HMI tags "AO"
   "DB332_AO_AO{1}_bRoZB1" : Byte = PLC DB332_AO.AO[1].bRoZB1, 1 s
   "DB332_AO_AO{1}_bSym" : Word = PLC DB332_AO.AO[1].bSym AT %DB1.DBB0, 1 s
   "DB332_AO_AO{1}_bSt_Tryb" : Word = PLC DB332_AO.AO[1].bSt_Tryb AT %DB1.DBW0, 1 s
   "DB332_AO_AO{1}_bSt_Urz" : Int = PLC DB332_AO.AO[1].bSt_Urz, 1 s
   "DB332_AO_AO{1}_bTrP" : Int = PLC DB332_AO.AO[1].bTrP AT %DB1.DBW0, 1 s
   "DB332_AO_AO{1}_yCzZadFiltru" : Byte = PLC DB332_AO.AO[1].yCzZadFiltru AT %DB1.DBW0, 1 s
   "DB332_AO_AO{1}_bB" : Byte = PLC DB332_AO.AO[1].bB AT %DB1.DBW0, 1 s
   "DB332_AO_AO{1}_rZH" : Real = PLC DB332_AO.AO[1].rZH AT %DB1.DBB0, 1 s
   "DB332_AO_AO{Nr}_rZL" : Real = PLC DB332_AO.AO[1].rZL AT %DB1.DBD0, 1 s
   "DB332_AO_AO{Nr}_rGHH" : Real = PLC DB332_AO.AO[1].rGHH AT %DB1.DBD0, 1 s
   "DB332_AO_AO{Nr}_rGH" : Real = PLC DB332_AO.AO[1].rGH AT %DB1.DBD0, 1 s
   "DB332_AO_AO{Nr}_rGL" : Real = PLC DB332_AO.AO[1].rGL AT %DB1.DBD0, 1 s
   "DB332_AO_AO{Nr}_rGLL" : Real = PLC DB332_AO.AO[1].rGLL AT %DB1.DBD0, 1 s
   "DB332_AO_AO{Nr}_rHI_LIM" : Real = PLC DB332_AO.AO[1].rHI_LIM, 1 s
   "DB332_AO_AO{Nr}_rRoManSter" : Real = PLC DB332_AO.AO[1].rRoManSter, 1 s
   "DB332_AO_AO{Nr}_rWy" : Real = PLC DB332_AO.AO[1].rWy, 1 s

HMI tags "DIO"
   "DB321_DIO_DIO{Nr}_bRoZB1" : Byte = PLC DB321_DIO.DIO[1].bRoZB1, 1 s
   "DB321_DIO_DIO{Nr}_bSt_Tryb" : Word = PLC DB321_DIO.DIO[1].bSt_Tryb AT %DB1.DBB0, 1 s
   "DB321_DIO_DIO{Nr}_bWySter" : Bool = PLC DB321_DIO.DIO[1].bWySter AT %DB1.DBW0, 1 s
   "DB321_DIO_DIO{Nr}_yCzZadOpzZal" : DWord = PLC DB321_DIO.DIO[1].yCzZadOpzZal AT %DB1.DBX0.0, 1 s
   "DB321_DIO_DIO{Nr}_yCzZadOpzWyl" : DWord = PLC DB321_DIO.DIO[1].yCzZadOpzWyl AT %DB1.DBD0, 1 s

HMI tags "DM"
   "DB323_DM1_DM1{Nr}_bRoZB1" : Byte = PLC DB323_DM1.DM1[1].bRoZB1, 1 s
   "DB323_DM1_DM1{Nr}_bRoZB2" : Byte = PLC DB323_DM1.DM1[1].bRoZB2 AT %DB1.DBB0, 1 s
   "DB323_DM1_DM1{Nr}_bSym" : Word = PLC DB323_DM1.DM1[1].bSym AT %DB1.DBB0, 1 s
   "DB323_DM1_DM1{Nr}_bSt_Tryb" : Word = PLC DB323_DM1.DM1[1].bSt_Tryb AT %DB1.DBW0, 1 s
   "DB323_DM1_DM1{Nr}_bSt_Urz" : Int = PLC DB323_DM1.DM1[1].bSt_Urz AT %DB1.DBW0, 1 s
   "DB323_DM1_DM1{Nr}_bTrP" : Int = PLC DB323_DM1.DM1[1].bTrP AT %DB1.DBW0, 1 s
   "DB323_DM1_DM1{Nr}_yCzZadOpzZal" : DWord = PLC DB323_DM1.DM1[1].yCzZadOpzZal AT %DB1.DBW0, 1 s
   "DB323_DM1_DM1{Nr}_yCzZadOpzWyl" : DWord = PLC DB323_DM1.DM1[1].yCzZadOpzWyl AT %DB1.DBD0, 1 s
   "DB323_DM1_DM1{1}" : UDT323_DM1 = PLC DB323_DM1.DM1[1] AT %DB1.DBB0, 1 s
   "DB323_DM1_DM1{2}" : UDT323_DM1 = PLC DB323_DM1.DM1[2] AT %DB1.DBW0, 1 s
   "DB323_DM1_DM1{3}" : UDT323_DM1 = PLC DB323_DM1.DM1[3] AT %DB1.DBW0, 1 s
   "DB323_DM1_DM1{4}" : UDT323_DM1 = PLC DB323_DM1.DM1[4] AT %DB1.DBW0, 1 s
   "DB323_DM1_DM1{5}" : UDT323_DM1 = PLC DB323_DM1.DM1[5] AT %DB1.DBW0, 1 s
   "DB323_DM1_DM1{Nr}_yCzZadOpzAlm" : Byte = PLC DB323_DM1.DM1[1].yCzZadOpzAlm AT %DB1.DBD0, 1 s
   "DB323_DM1_DM1{Nr}_bWySter" : Bool = PLC DB323_DM1.DM1[1].bWySter AT %DB1.DBD0, 1 s

HMI tags "DV"
   "DB322_DV1_DV1{Nr}_bRoZB1" : Byte = PLC DB322_DV1.DV1[1].bRoZB1, 1 s
   "DB322_DV1_DV1{Nr}_bRoZB2" : Byte = PLC DB322_DV1.DV1[1].bRoZB2 AT %DB1.DBB0, 1 s
   "DB322_DV1_DV1{Nr}_bSym" : Word = PLC DB322_DV1.DV1[1].bSym AT %DB1.DBB0, 1 s
   "DB322_DV1_DV1{Nr}_bSt_Tryb" : Word = PLC DB322_DV1.DV1[1].bSt_Tryb AT %DB1.DBW0, 1 s
   "DB322_DV1_DV1{Nr}_bSt_Urz" : Int = PLC DB322_DV1.DV1[1].bSt_Urz AT %DB1.DBW0, 1 s
   "DB322_DV1_DV1{Nr}_bTrP" : Int = PLC DB322_DV1.DV1[1].bTrP AT %DB1.DBW0, 1 s
   "DB322_DV1_DV1{Nr}_yCzZadOpzZal" : DWord = PLC DB322_DV1.DV1[1].yCzZadOpzZal AT %DB1.DBW0, 1 s
   "DB322_DV1_DV1{Nr}_yCzZadOpzWyl" : DWord = PLC DB322_DV1.DV1[1].yCzZadOpzWyl, 1 s
   "DB322_DV1_DV1{Nr}_yCzZadOpzAlm" : Byte = PLC DB322_DV1.DV1[1].yCzZadOpzAlm AT %DB1.DBD0, 1 s
   "DB322_DV1_DV1{1}" : UDT322_DVI = PLC DB322_DV1.DV1[1] AT %DB1.DBD0, 1 s
   "DB322_DV1_DV1{2}" : UDT322_DVI = PLC DB322_DV1.DV1[2] AT %DB1.DBW0, 1 s
   "DB322_DV1_DV1{Nr}_bWySter" : Bool = PLC DB322_DV1.DV1[1].bWySter AT %DB1.DBD0, 1 s

HMI tags "Tag table_1"
   "DB_DM_pump1Tank1out_inTurnOnDelay" : DInt = PLC DB_DM.pump1Tank1out.inTurnOnDelay, 1 s
   "DB_DM_pump1Tank1out_inTurnOffDelay" : DInt = PLC DB_DM.pump1Tank1out.inTurnOffDelay, 1 s
   "DB_DM_pump1Tank1out_inAlarmDelay" : DInt = PLC DB_DM.pump1Tank1out.inAlarmDelay, 1 s
   "DB_DM_pump1Tank1out_oFaultCode" : Byte = PLC DB_DM.pump1Tank1out.oFaultCode, 1 s
   "DB_DM_pump1Tank1out_oStatusCode" : Word = PLC DB_DM.pump1Tank1out.oStatusCode, 1 s
   "DB_DM_pump1Tank1out_oStatus" : Int = PLC DB_DM.pump1Tank1out.oStatus, 1 s
   "DB_DM_pump1Tank1out_oControlMode" : Int = PLC DB_DM.pump1Tank1out.oControlMode, 1 s
   "DB_DM_pump1Tank1out_inCmdOper" : Word = PLC DB_DM.pump1Tank1out.inCmdOper, 1 s
   "DB_DM_pump1Tank1out_inSimOper" : Word = PLC DB_DM.pump1Tank1out.inSimOper, 1 s
   "DB_DM_pump1Tank1out_inCmdOperImp" : Word = PLC DB_DM.pump1Tank1out.inCmdOperImp, 1 s
   "DB_DM_pump2Tank1in_inTurnOnDelay" : DInt = PLC DB_DM.pump2Tank1in.inTurnOnDelay, 1 s
   "DB_DM_pump2Tank1in_inTurnOffDelay" : DInt = PLC DB_DM.pump2Tank1in.inTurnOffDelay, 1 s
   "DB_DM_pump2Tank1in_inAlarmDelay" : DInt = PLC DB_DM.pump2Tank1in.inAlarmDelay, 1 s
   "DB_DM_pump2Tank1in_oFaultCode" : Byte = PLC DB_DM.pump2Tank1in.oFaultCode, 1 s
   "DB_DM_pump2Tank1in_oStatusCode" : Word = PLC DB_DM.pump2Tank1in.oStatusCode, 1 s
   "DB_DM_pump2Tank1in_oStatus" : Int = PLC DB_DM.pump2Tank1in.oStatus, 1 s
   "DB_DM_pump2Tank1in_oControlMode" : Int = PLC DB_DM.pump2Tank1in.oControlMode, 1 s
   "DB_DM_pump2Tank1in_inCmdOper" : Word = PLC DB_DM.pump2Tank1in.inCmdOper, 1 s
   "DB_DM_pump2Tank1in_inSimOper" : Word = PLC DB_DM.pump2Tank1in.inSimOper, 1 s
   "DB_DM_pump2Tank1in_inCmdOperImp" : Word = PLC DB_DM.pump2Tank1in.inCmdOperImp, 1 s

text list "DMI_Obiekt": 0 '1. Naped mostu / M321'; 1 '2. Naped wozka / M123'; 2 '3. Pompa chwytaka'; 3 '4. Naped wciagarki'; 4 '5. Naped zwijaka'

text list "AO_Obiekt": 0 'AO1'; 1 'AO2'

text list "DIO_Obiekt": 0 '1. DI_Przek_Bezp / B231'; 1 '2. DI_Stop / dd'; 2 '3. DI_Start'; 3 '4. DI_Deblokada'; 4 '5. DI_Podoszenie'; 5 '6. DI_Opuszczanie'; 6 '7. DI_Otw_Chwyt'; 7 '8. DI_Zamkn_Chwyt'; 8 '9. DI_Wozek_Prawo'; 9 '10. DI_Wozek_Lewo'; 10 '11. DI_Most_Przod'; 11 '12. DI_Most_Tyl'; 12 '13. DI_Kranc_Podn'; 13 '14. DI_Kranc_Opuszcz'; 14 '15. DI_Kranc_Lina'; 15 '16. DI_Kranc_Potw_Zamkn_Hamul'; 16 '17. DI_Zabezp_Hamul_Podn'; 17 '18. DI_Blad_Fal_Podn'; 18 '19. DI_Zabezp_Term_Siln_Podn'; 19 '20. DI_Kranc_Wozek_Lewo_Zatrzym'; 20 '21. DI_Kranc_Wozek_Lewo_Zwoln'; 21 '22. DI_Kranc_Wozek_Prawo_Zatrzym'; 22 '23. DI_Kranc_Wozek_Prawo_Zwoln'; 23 '24. DI_Czujn_Ustal_Wozek'; 24 '25. DI_Zabezp_Hamul_Wozek'; 25 '26. DI_Blad_Fal_Wozek'; 26 '27. DI_Zabezp_PTC_M301_Wozek'; 27 '28. DI_Zabezp_PTC_M302_Wozek'; 28 '29. DI_Kranc_Most_Przod_Zatrzym'; 29 '30. DI_Kranc_Most_Przod_Zwoln'; 30 '31. DI_Kranc_Most_Tyl_Zatrzym'; 31 '32. DI_Kranc_Most_Tyl_Zwoln'; 32 '33. DI_Czujn_Ustal_Most'; 33 '34. DI_Zabezp_Hamul_Most'; 34 '35. DI_Blad_Fal_Most'; 35 '36. DI_Zabezp_Term_Siln1_Most'; 36 '37. DI_Zabezp_Term_Siln2_Most'; 37 '38. DI_Zabezp_Zwijak'; 38 '39. DI_Blad_Zasil_Obw_Analog'; 39 '40. DI_Zabezp_Siln_Chwyt_M801'; 40 '41. DI_Zabezp_Obw_Ster_Chwyt'; 41 '42. DI_Zabezp_Term_Siln_Chwyt'; 42 '43. DI_Kranc_Otw_Chwy'; 43 '44. DI_Kranc_Zamkn_Chwyt'; 44 '45. DI_Rezerwa'; 45 '46. DI_Czujn_Przechyl_Chwyt'; 46 '47. DI_Czujn_Poziom_Oleju'; 47 '48. DI_Czujn_Temp_Oleju'; 48 '49. DI_Kontrol_Zasil_Chwyt'; 49 '50. DI_Chwyt_Podlaczony'; 50 '51. DI_Przel_Ster_Radiowe'; 51 '52. DI_Zalacz_Suwnice'; 52 '53. DI_Wylacz_Suwnice'; 53 '54. DI_Zuzyc_Tarczy_Hamul'; 54 '55. DI_Kranc_Otw_Hamul'; 69 '70. DO_Start'; 70 '71. DO_Syrena'; 71 '72. DO_Podnoszenie'; 72 '73. DO_Opuszczanie'; 73 '74. DO_Awr_Podn'; 74 '75. DO_Potw_Hamul'; 75 '76. DO_Przciaz'; 76 '77. DO_Wozek_Lewo'; 77 '78. DO_Wozek_Prawo'; 78 '79. DO_Awr_Wozek'; 79 '80. DO_Most_Przod'; 80 '81. DO_Most_Tyl'; 81 '82. DO_Awr_Most'; 82 '83. DO_Zal_Zwijak'; 83 '84. DO_Awr_Zwijak'; 84 '85. DO_Lina_PozaRowiem'; 85 '86. DO_Otw_Chwytak'; 86 '87. DO_Zamkn_Chwytak'; 87 '88. DO_Blad_Chwytak'; 88 '89. DO_Zabezp_PompChytak'; 89 '90. DO_Zalacz_Skaner'; 90 '91. DO_Went_Szafa'

text list "AI_Obiekt": 0 'AI1'; 1 'AI2'

text list "Awaria": 0 'BRAK AWARII'; 1 'AWARIA!'; 2..32 'BRAK AWARII'

text list "DMI_Status": 1 'Wyłącznik Remontowy'; 2 'Sterowanie Lokalne'; 4 'Tryb Manualny'; 8 'Tryb Automatyczny'

text list "DV1_Status": 1 'Wyłącznik Remontowy'; 2 'Sterowanie Lokalne'; 4 'Tryb Manualny'; 8 'Tryb Automatyczny'

text list "DVI_Obiekt": 0 '1. Chwytak otwarcie / Z456'; 1 '2. Chwytak zamkniecie / Z456'

Template "Template_1" 1280x800
   Button "Exit" at 1182,752 size 67x47; TextOff 'Exit'; PictureOff "ExitRuntime_KTP1200_Basic_PN_TR"; PictureOn "ExitRuntime_KTP1200_Basic_PN_TR"
      on Release: StopRuntime(0)
   Button "Template_Button" at 1054,752 size 67x47; TextOff 'Text'
   Button "Template_Button_1" at 926,752 size 67x47; TextOff 'Text'
   Button "Template_Button_2" at 798,752 size 67x47; TextOff 'Text'
   Button "Template_Button_3" at 670,752 size 67x47; TextOff 'Text'
   Button "Template_Button_4" at 542,752 size 67x47; TextOff 'Text'
   Button "Template_Button_5" at 414,752 size 67x47; TextOff 'Text'
   Button "Template_Button_6" at 286,752 size 67x47; TextOff 'Text'
   Button "Alarms" at 158,752 size 67x47; TextOff 'Alarms'; PictureOff "AlarmDisplay_KTP1200_Basic_PN_TR"; PictureOn "AlarmDisplay_KTP1200_Basic_PN_TR"
      on Release: function_ef3f5d25("Alarm window_Unacknowledged", -1)
   Button "Start screen" at 30,752 size 67x47; TextOff 'Start screen'; PictureOff "NavigateHome_KTP1200_Basic_PN_TR"; PictureOn "NavigateHome_KTP1200_Basic_PN_TR"
      on Release: ActivateScreen("Root screen", 0)
   SymbolicIOField "Symbolic_IO_Field_Screen" at 87,9 size 1086x30; TextOff '0'; TextOn '1'; TextList "TextList_ScreenNames"
      ProcessValue <- "Tag_ScreenNumber"
      on Change: ActivateScreenByNumber("Tag_ScreenNumber", 0)
   DateTimeField "HmiScreenItemData" at 1175,24 size 105x24
   DateTimeField "HmiScreenItemData_1" at 1175,0 size 105x24
   GraphicView "Logo" at 0,0 size 85x48; Picture "Logo of HMI_1"

screen "Root screen" 1280x800, template "Template_1"
   on GenerateScreen: SetTag("Tag_ScreenNumber", 1)
   Button "HmiScreenItemData" at 36,84 size 159x47; TextOff 'Screen0'; PictureOff "Navigates to Screen0 for KTP1200 Basic+ PN 17.0.0.0"; PictureOn "Navigates to Screen0 for KTP1200 Basic+ PN 17.0.0.0"
      on Release: ActivateScreen("Screen0", 0)

screen "Screen0" 1280x800, template "Template_1"
   on GenerateScreen: SetTag("Tag_ScreenNumber", 2)
   TextField "HmiScreenItemData" at 128,384 size 1024x27; Text 'Screen0'
   Button "Back" at 1,49 size 159x47; TextOff 'Back'
      on Release: ActivateScreen("Root screen", 0)

screen "Service" 1280x800, template "Template_1"
   on GenerateScreen: SetTag("Tag_ScreenNumber", 10)
   TextField "Text field_1" at 560,183 size 163x25; Text 'Zakres pomiarowy'
   TextField "Text field_2" at 543,217 size 57x25; Text 'Górny'
   TextField "Text field_3" at 545,259 size 55x25; Text 'Dolny'
   TextField "Text field_4" at 573,301 size 132x25; Text 'Tryb manualny'
   TextField "Text field_5" at 530,432 size 108x25; Text 'Progi alarm.'
   TextField "Text field_6" at 642,431 size 101x25; Text 'Blok. alarm'
   TextField "Text field_7" at 560,103 size 174x25; Text 'Wejścia analogowe / Pomiary analogowe'
   SymbolicIOField "Symbolic I/O field_1" at 536,138 size 222x31; TextOn '1'; TextOff '0'; TextList "AI_Obiekt"
      ProcessValue <- "Nr_AI"
   IOField "I/O field_3" at 627,212 size 110x35; FormatPattern s999.9
      ProcessValue <- "DB331_AI_AI{Nr}_rZH"
   IOField "I/O field_4" at 627,255 size 110x35; FormatPattern s999.9
      ProcessValue <- "DB331_AI_AI{Nr}_rZL"
   Button "Button_5" at 534,331 size 97x35; TextOn 'Wyłączony'; TextOff 'ON / Wyłączony'
      on Click: function_a9b64e44("DB331_AI_AI{Nr}_bRoZB1", 3); function_b3f726e6("DB331_AI_AI{Nr}_bRoZB1", 0)
      Appearance <- "DB331_AI_AI{Nr}_bRoZB1"
   IOField "I/O field_5" at 584,374 size 110x35; FormatPattern s999.9
      Appearance <- "DB331_AI_AI{Nr}_bRoZB1"
      ProcessValue <- "DB331_AI_AI{Nr}_rRoManSter"
   IOField "I/O field_6" at 533,463 size 96x32; FormatPattern 999.9
      ProcessValue <- "DB331_AI_AI{Nr}_rGHH"
   Button "Button_7" at 695,463 size 54x33; TextOn 'OFF'; TextOff 'OFF'
      on Click: function_a9b64e44("DB331_AI_AI{Nr}_bB", 0)
      Appearance <- "DB331_AI_AI{Nr}_bB"
   IOField "I/O field_7" at 533,515 size 96x32; FormatPattern 999.9
      ProcessValue <- "DB331_AI_AI{Nr}_rGH"
   IOField "I/O field_8" at 533,567 size 96x32; FormatPattern 999.9
      ProcessValue <- "DB331_AI_AI{Nr}_rGL"
   IOField "I/O field_9" at 533,620 size 96x32; FormatPattern 999.9
      ProcessValue <- "DB331_AI_AI{Nr}_rGLL"
   Button "Button_9" at 695,516 size 54x33; TextOn 'OFF'; TextOff 'OFF'
      on Click: function_a9b64e44("DB331_AI_AI{Nr}_bB", 0)
      Appearance <- "DB331_AI_AI{Nr}_bB"
   Button "Button_11" at 695,568 size 54x33; TextOn 'OFF'; TextOff 'OFF'
      on Click: function_a9b64e44("DB331_AI_AI{Nr}_bB", 0)
      Appearance <- "DB331_AI_AI{Nr}_bB"
   Button "Button_13" at 695,621 size 54x33; TextOn 'OFF'; TextOff 'OFF'
      on Click: function_a9b64e44("DB331_AI_AI{Nr}_bB", 0)
      Appearance <- "DB331_AI_AI{Nr}_bB"
   Button "Button_4" at 651,331 size 97x35; TextOn 'Włączony'; TextOff 'OFF / Włączony'
      on Click: function_b3f726e6("DB331_AI_AI{Nr}_bRoZB1", 3); function_a9b64e44("DB331_AI_AI{Nr}_bRoZB1", 0)
      Appearance <- "DB331_AI_AI{Nr}_bRoZB1"
   Button "Button_6" at 642,463 size 54x33; TextOn 'ON'; TextOff 'ON'
      on Click: function_b3f726e6("DB331_AI_AI{Nr}_bB", 0)
      Appearance <- "DB331_AI_AI{Nr}_bB"
   Button "Button_8" at 642,516 size 54x33; TextOn 'ON'; TextOff 'ON'
      on Click: function_a9b64e44("DB331_AI_AI{Nr}_bB", 0)
      Appearance <- "DB331_AI_AI{Nr}_bB"
   Button "Button_10" at 642,568 size 54x33; TextOn 'ON'; TextOff 'ON'
      on Click: function_a9b64e44("DB331_AI_AI{Nr}_bB", 0)
      Appearance <- "DB331_AI_AI{Nr}_bB"
   Button "Button_12" at 642,621 size 54x33; TextOn 'ON'; TextOff 'ON'
      on Click: function_a9b64e44("DB331_AI_AI{Nr}_bB", 0)
      Appearance <- "DB331_AI_AI{Nr}_bB"
   TextField "Text field_8" at 226,246 size 132x25; Text 'Tryb manualny'
   TextField "Text field_9" at 207,312 size 170x25; Text 'Sterowanie manual / Sterowanie'
   Circle "Circle_1" at 275,206 size 30x30
      Appearance <- "DB321_DIO_DIO{Nr}_bWySter"
   TextField "Text field_10" at 220,178 size 147x25; Text 'Wejście/Wyjście'
   TextField "Text field_12" at 193,455 size 200x42; Text 'Zad. czas opóźn. załącz. Zadany czas opóźnienia załączenia'
   TextField "Text field_13" at 92,102 size 221x25; Text 'Wejścia/Wyjścia cyfrowe'
   Button "Button_14" at 191,271 size 97x35; TextOn 'ON'; TextOff 'ON'
      on Click: function_a9b64e44("DB321_DIO_DIO{Nr}_bRoZB1", 0)
      Appearance <- "DB321_DIO_DIO{Nr}_bRoZB1"
   Button "Button_16" at 191,336 size 97x35; TextOn 'Aktywne'; TextOff 'ON / Aktywne'
      on Click: function_b3f726e6("DB321_DIO_DIO{Nr}_bRoZB1", 3)
      Appearance <- "DB321_DIO_DIO{Nr}_bRoZB1"
      ObjectEnable <- "DB321_DIO.DIO[Nr].bRoZB1"
   IOField "I/O field_2" at 242,551 size 96x32; FormatPattern 999
      ProcessValue <- "DB321_DIO_DIO{Nr}_yCzZadOpzWyl"
   IOField "I/O field_1" at 242,490 size 96x32; FormatPattern 999
      ProcessValue <- "DB321_DIO_DIO{Nr}_yCzZadOpzZal"
   Button "Button_1" at 300,271 size 97x35; TextOn 'OFF'; TextOff 'OFF'
      on Click: function_b3f726e6("DB321_DIO_DIO{Nr}_bRoZB1", 0)
      Appearance <- "DB321_DIO_DIO{Nr}_bRoZB1"
   Button "Button_3" at 300,336 size 97x35; TextOn 'Nieaktywne'; TextOff 'OFF / Nieaktywne'
      on Click: function_a9b64e44("DB321_DIO_DIO{Nr}_bRoZB1", 3)
      Appearance <- "DB321_DIO_DIO{Nr}_bRoZB1"
      ObjectEnable <- "DB321_DIO.DIO[Nr].bRoZB1"
   SymbolicIOField "Symbolic I/O field_2" at 100,138 size 390x31; TextOn '1'; TextOff '0'; TextList "DIO_Obiekt"
      ProcessValue <- "Nr_DIO"
   TextField "Text field_14" at 905,179 size 183x25; Text 'Granica skal. wyjścia'
   TextField "Text field_15" at 932,247 size 132x25; Text 'Tryb manualny'
   TextField "Text field_16" at 915,104 size 170x25; Text 'Wyjścia analogowe'
   IOField "I/O field_10" at 945,205 size 110x35; FormatPattern s999.9
      ProcessValue <- "DB332_AO_AO{Nr}_rHI_LIM"
   Button "Button_2" at 998,272 size 97x35; TextOn 'OFF'; TextOff 'OFF'
      on Click: function_a9b64e44("DB332_AO_AO{1}_bRoZB1", 3); function_b3f726e6("DB332_AO_AO{1}_bRoZB1", 0)
      Appearance <- "DB332_AO_AO{1}_bRoZB1"
   Button "Button_15" at 900,272 size 97x35; TextOn 'ON'; TextOff 'ON'
      on Click: function_b3f726e6("DB332_AO_AO{1}_bRoZB1", 3); function_a9b64e44("DB332_AO_AO{1}_bRoZB1", 0)
      Appearance <- "DB332_AO_AO{1}_bRoZB1"
   IOField "I/O field_11" at 942,316 size 110x35; FormatPattern s999.9
      Appearance <- "DB332_AO_AO{1}_bRoZB1"
      ProcessValue <- "DB332_AO_AO{Nr}_rRoManSter"
   SymbolicIOField "Symbolic I/O field_3" at 898,137 size 204x31; TextOn '1'; TextOff '0'; TextList "AO_Obiekt"
      ProcessValue <- "Nr_AO"
   TextField "Text field_24" at 190,516 size 204x42; Text 'Zad. czas opóźn. wyłącz. Zadany czas opóźnienia załączenia'
   Button "Button_17" at 1069,671 size 188x32; TextOn 'Zawory i silniki'; TextOff 'Zawory i silniki'
      on Click: ActivateScreen("Service2", 0)
   GraphicView "Graphic view_11" at 1222,672 size 36x30; Picture "Graphic_97"
   TextField "Text field_36" at 214,383 size 156x25; Text 'Praca z wyjściami / Sterowanie'
   Button "Button_18" at 191,410 size 97x35; TextOn 'ON'; TextOff 'ON'
      on Click: function_b3f726e6("DB321_DIO_DIO{Nr}_bRoZB1", 2)
      ObjectEnable <- "DB322_DV1.DV1[Nr].bRoZB1"
      Appearance <- "DB321_DIO_DIO{Nr}_bRoZB1"
   Button "Button_19" at 300,410 size 97x35; TextOn 'OFF'; TextOff 'OFF'
      on Click: function_a9b64e44("DB321_DIO_DIO{Nr}_bRoZB1", 2)
      ObjectEnable <- "DB322_DV1.DV1[Nr].bRoZB1"
      Appearance <- "DB321_DIO_DIO{Nr}_bRoZB1"
   Button "Button_20" at 900,445 size 188x32; TextOn 'Zawory i silniki'; TextOff 'Włacz symulacje / Zawory i silniki'

screen "Service2" 1280x800, template "Template_1"
   on GenerateScreen: SetTag("Tag_ScreenNumber", 12)
   TextField "Text field_17" at 364,324 size 188x22; Text 'Zad. czas opóźn. wyłącz:'
   TextField "Text field_18" at 371,266 size 174x22; Text 'Zad. czas opóź. załącz:'
   TextField "Text field_19" at 373,382 size 173x22; Text 'Zad. czas monitoringu:'
   TextField "Text field_20" at 365,511 size 185x23; Text 'Monitoring potwierdz.'
   TextField "Text field_21" at 368,448 size 180x23; Text 'Symulacja potwierdz.'
   TextField "Text field_22" at 366,208 size 142x22; Text 'Zawór zamknięty / Potwierdz. załącz.'
   TextField "Text field_23" at 366,237 size 147x22; Text 'Zawór otwarty / Potwierdz. wyłącz.'
   TextField "Text field_11" at 314,110 size 69x25; Text 'Zawory'
   TextField "Text field_25" at 169,446 size 132x25; Text 'Tryb manualny'
   TextField "Text field_26" at 201,242 size 84x22; Text 'INTERLOK'
      Appearance <- "DB322_DV1_DV1{Nr}_bSt_Tryb"
   SymbolicIOField "Symbolic I/O field_4" at 139,208 size 205x32; TextOn '1'; TextOff '0'; TextList "DV1_Status"
      ProcessValue <- "DB322_DV1_DV1{Nr}_bTrP"
      Appearance <- "DB322_DV1_DV1{Nr}_bTrP"
   TextField "Text field_29" at 198,183 size 95x25; Text 'Tryb Pracy'
   TextField "Text field_30" at 187,510 size 102x25; Text 'Sterowanie'
   TextField "Text field_31" at 393,183 size 127x25; Text 'Potwierdzenia'
   TextField "Text field_27" at 174,265 size 135x25; Text 'Obsługa Awarii'
   SymbolicIOField "Symbolic I/O field_6" at 177,292 size 130x32; TextOn '1'; TextOff '0'; TextList "Awaria"
      ProcessValue <- "DB322_DV1_DV1{Nr}_bSt_Urz"
      Appearance <- "DB322_DV1_DV1{Nr}_bSt_Urz"
   TextField "Text field_28" at 148,370 size 184x22; Text 'BŁĄD POTWIERDZENIA'
      Appearance <- "DB322_DV1_DV1{Nr}_bSt_Tryb"
   TextField "Text field_32" at 148,395 size 184x22; Text 'BRAK GOTOWOŚCI'
      Appearance <- "DB322_DV1_DV1{Nr}_bSt_Tryb"
   TextField "Text field_33" at 148,419 size 184x22; Text 'AWARIA ZEWNĘTRZNA'
      Appearance <- "DB322_DV1_DV1{Nr}_bSt_Tryb"
   TextField "Text field_8" at 896,110 size 57x25; Text 'Silniki'
   Button "Button_20" at 355,536 size 97x32; TextOn 'ON'; TextOff 'ON'
      on Click: function_b3f726e6("DB322_DV1_DV1{Nr}_bRoZB1", 6)
      Appearance <- "DB322_DV1_DV1{Nr}_bRoZB1"
   Button "Button_21" at 462,536 size 97x32; TextOn 'OFF'; TextOff 'OFF'
      on Click: function_a9b64e44("DB322_DV1_DV1{Nr}_bRoZB1", 6)
      Appearance <- "DB322_DV1_DV1{Nr}_bRoZB1"
   Button "Button_22" at 355,474 size 97x32; TextOn 'ON'; TextOff 'ON'
      on Click: function_b3f726e6("DB322_DV1_DV1{Nr}_bRoZB1", 1)
      Appearance <- "DB322_DV1_DV1{Nr}_bRoZB1"
   Button "Button_23" at 462,474 size 97x32; TextOn 'OFF'; TextOff 'OFF'
      on Click: function_a9b64e44("DB322_DV1_DV1{Nr}_bRoZB1", 1)
      Appearance <- "DB322_DV1_DV1{Nr}_bRoZB1"
   IOField "I/O field_12" at 411,291 size 96x32; FormatPattern 999
      ProcessValue <- "DB322_DV1_DV1{Nr}_yCzZadOpzZal"
   IOField "I/O field_13" at 411,349 size 96x32; FormatPattern 999
      ProcessValue <- "DB322_DV1_DV1{Nr}_yCzZadOpzWyl"
   IOField "I/O field_14" at 411,407 size 96x32; FormatPattern 999
      ProcessValue <- "DB322_DV1_DV1{Nr}_yCzZadOpzAlm"
   Button "Button_17" at 138,472 size 97x35; TextOn 'ON'; TextOff 'ON'
      on Click: function_a9b64e44("DB322_DV1_DV1{Nr}_bRoZB1", 0)
      Appearance <- "DB322_DV1_DV1{Nr}_bRoZB1"
   Button "Button_18" at 245,472 size 97x35; TextOn 'OFF'; TextOff 'OFF'
      on Click: function_b3f726e6("DB322_DV1_DV1{Nr}_bRoZB1", 0)
      Appearance <- "DB322_DV1_DV1{Nr}_bRoZB1"
   Button "Button_19" at 137,534 size 97x35; TextOn 'ON'; TextOff 'ON'
      on Click: function_b3f726e6("DB322_DV1_DV1{Nr}_bRoZB1", 3)
      ObjectEnable <- "DB322_DV1.DV1[Nr].bRoZB1"
      Appearance <- "DB322_DV1_DV1{Nr}_bRoZB1"
   Button "Button_24" at 245,534 size 97x35; TextOn 'OFF'; TextOff 'OFF'
      on Click: function_a9b64e44("DB322_DV1_DV1{Nr}_bRoZB1", 3)
      ObjectEnable <- "DB322_DV1.DV1[Nr].bRoZB1"
      Appearance <- "DB322_DV1_DV1{Nr}_bRoZB1"
   SymbolicIOField "Symbolic I/O field_5" at 247,146 size 204x31; TextOn '1'; TextOff '0'; TextList "DVI_Obiekt"
      ProcessValue <- "Nr_DV"
   Button "Button_25" at 189,329 size 110x35; TextOn 'Reset Awarii'; TextOff 'Reset Awarii'
      on Click: function_b3f726e6("DB322_DV1_DV1{Nr}_bRoZB2", 0)
   TextField "Text field_1" at 939,324 size 188x22; Text 'Zad. czas opóźn. wyłącz:'
   TextField "Text field_2" at 946,266 size 174x22; Text 'Zad. czas opóź. załącz:'
   TextField "Text field_3" at 948,382 size 173x22; Text 'Zad. czas monitoringu:'
   TextField "Text field_4" at 940,511 size 185x23; Text 'Monitoring potwierdz.'
   TextField "Text field_5" at 943,448 size 180x23; Text 'Symulacja potwierdz.'
   TextField "Text field_6" at 941,208 size 142x22; Text 'Potwierdz. załącz.'
   TextField "Text field_7" at 941,237 size 147x22; Text 'Potwierdz. wyłącz.'
   Circle "Circle_1" at 1092,207 size 25x25
      Appearance <- "DB323_DM1_DM1{Nr}_bSt_Urz"
   Circle "Circle_4" at 1092,237 size 25x25
      Appearance <- "DB323_DM1_DM1{Nr}_bSt_Urz"
   TextField "Text field_9" at 744,446 size 132x25; Text 'Tryb manualny'
   TextField "Text field_10" at 776,242 size 84x22; Text 'INTERLOK'
      Appearance <- "DB323_DM1_DM1{Nr}_bSt_Tryb"
   SymbolicIOField "Symbolic I/O field_1" at 714,208 size 205x32; TextOn '1'; TextOff '0'; TextList "DMI_Status"
      ProcessValue <- "DB323_DM1_DM1{Nr}_bTrP"
      Appearance <- "DB323_DM1_DM1{Nr}_bTrP"
   TextField "Text field_12" at 773,183 size 95x25; Text 'Tryb Pracy'
   TextField "Text field_13" at 762,510 size 102x25; Text 'Sterowanie'
   TextField "Text field_14" at 968,183 size 127x25; Text 'Potwierdzenia'
   TextField "Text field_15" at 749,265 size 135x25; Text 'Obsługa Awarii'
   SymbolicIOField "Symbolic I/O field_2" at 752,292 size 130x32; TextOn '1'; TextOff '0'; TextList "Awaria"
      ProcessValue <- "DB323_DM1_DM1{Nr}_bSt_Urz"
      Appearance <- "DB323_DM1_DM1{Nr}_bSt_Urz"
   TextField "Text field_16" at 723,370 size 184x22; Text 'BŁĄD POTWIERDZENIA'
      Appearance <- "DB323_DM1_DM1{Nr}_bSt_Tryb"
   TextField "Text field_24" at 723,395 size 184x22; Text 'BRAK GOTOWOŚCI'
      Appearance <- "DB323_DM1_DM1{Nr}_bSt_Tryb"
   TextField "Text field_34" at 723,419 size 184x22; Text 'AWARIA ZEWNĘTRZNA'
      Appearance <- "DB323_DM1_DM1{Nr}_bSt_Tryb"
   Button "Button_1" at 930,536 size 97x32; TextOn 'ON'; TextOff 'ON'
      on Click: function_b3f726e6("DB323_DM1_DM1{Nr}_bRoZB1", 6)
      Appearance <- "DB323_DM1_DM1{Nr}_bRoZB1"
   Button "Button_2" at 1037,536 size 97x32; TextOn 'OFF'; TextOff 'OFF'
      on Click: function_a9b64e44("DB323_DM1_DM1{Nr}_bRoZB1", 6)
      Appearance <- "DB323_DM1_DM1{Nr}_bRoZB1"
   Button "Button_3" at 930,474 size 97x32; TextOn 'ON'; TextOff 'ON'
      on Click: function_b3f726e6("DB323_DM1_DM1{Nr}_bRoZB1", 1)
      Appearance <- "DB323_DM1_DM1{Nr}_bRoZB1"
   Button "Button_4" at 1037,474 size 97x32; TextOn 'OFF'; TextOff 'OFF'
      on Click: function_a9b64e44("DB323_DM1_DM1{Nr}_bRoZB1", 1)
      Appearance <- "DB323_DM1_DM1{Nr}_bRoZB1"
   IOField "I/O field_1" at 986,291 size 96x32; FormatPattern 999
      ProcessValue <- "DB323_DM1_DM1{Nr}_yCzZadOpzZal"
   IOField "I/O field_2" at 986,349 size 96x32; FormatPattern 999
      ProcessValue <- "DB323_DM1_DM1{Nr}_yCzZadOpzWyl"
   IOField "I/O field_3" at 986,407 size 96x32; FormatPattern 999
      ProcessValue <- "DB323_DM1_DM1{Nr}_yCzZadOpzAlm"
   Button "Button_5" at 713,472 size 97x35; TextOn 'ON'; TextOff 'ON'
      on Click: function_a9b64e44("DB323_DM1_DM1{Nr}_bRoZB1", 0)
      Appearance <- "DB323_DM1_DM1{Nr}_bRoZB1"
   Button "Button_6" at 820,472 size 97x35; TextOn 'OFF'; TextOff 'OFF'
      on Click: function_b3f726e6("DB323_DM1_DM1{Nr}_bRoZB1", 0)
      Appearance <- "DB323_DM1_DM1{Nr}_bRoZB1"
   Button "Button_7" at 712,534 size 97x35; TextOn 'ON'; TextOff 'ON'
      on Click: function_b3f726e6("DB323_DM1_DM1{Nr}_bRoZB1", 3)
      ObjectEnable <- "DB322_DV1.DV1[Nr].bRoZB1"
      Appearance <- "DB323_DM1_DM1{Nr}_bRoZB1"
   Button "Button_8" at 820,534 size 97x35; TextOn 'OFF'; TextOff 'OFF'
      on Click: function_a9b64e44("DB323_DM1_DM1{Nr}_bRoZB1", 3)
      ObjectEnable <- "DB322_DV1.DV1[Nr].bRoZB1"
      Appearance <- "DB323_DM1_DM1{Nr}_bRoZB1"
   SymbolicIOField "Symbolic I/O field_3" at 822,146 size 204x31; TextOn '1'; TextOff '0'; TextList "DMI_Obiekt"
      ProcessValue <- "Nr_DM"
   Button "Button_9" at 763,329 size 110x35; TextOn 'Reset Awarii'; TextOff 'Reset Awarii'
      on Click: function_b3f726e6("DB323_DM1_DM1{Nr}_bRoZB2", 0)
   TextField "Text field_35" at 773,572 size 102x25; Text 'Kierunek / Sterowanie'
   Button "Button_10" at 712,599 size 97x35; TextOn 'ON'; TextOff 'Lewo / ON'
      on Click: function_b3f726e6("DB323_DM1_DM1{Nr}_bRoZB1", 4)
      ObjectEnable <- "DB322_DV1.DV1[Nr].bRoZB1"
      Appearance <- "DB323_DM1_DM1{Nr}_bRoZB1"
   Button "Button_11" at 820,599 size 97x35; TextOn 'OFF'; TextOff 'Prawo / OFF'
      on Click: function_a9b64e44("DB323_DM1_DM1{Nr}_bRoZB1", 4)
      ObjectEnable <- "DB322_DV1.DV1[Nr].bRoZB1"
      Appearance <- "DB323_DM1_DM1{Nr}_bRoZB1"
   TextField "Text field_36" at 163,585 size 156x25; Text 'Praca z wyjściami / Sterowanie'
   Button "Button_12" at 137,611 size 97x35; TextOn 'ON'; TextOff 'ON'
      on Click: function_b3f726e6("DB322_DV1_DV1{Nr}_bRoZB1", 2)
      ObjectEnable <- "DB322_DV1.DV1[Nr].bRoZB1"
      Appearance <- "DB322_DV1_DV1{Nr}_bRoZB1"
   Button "Button_13" at 245,611 size 97x35; TextOn 'OFF'; TextOff 'OFF'
      on Click: function_a9b64e44("DB322_DV1_DV1{Nr}_bRoZB1", 2)
      ObjectEnable <- "DB322_DV1.DV1[Nr].bRoZB1"
      Appearance <- "DB322_DV1_DV1{Nr}_bRoZB1"
   TextField "Text field_37" at 390,585 size 126x25; Text 'Wyjście steruj / Sterowanie'
   Circle "Circle_5" at 437,614 size 30x30
      Appearance <- "DB322_DV1_DV1{Nr}_bWySter"
   TextField "Text field_38" at 738,651 size 156x25; Text 'Praca z wyjściami / Sterowanie'
   Button "Button_14" at 712,677 size 97x35; TextOn 'ON'; TextOff 'ON'
      on Click: function_b3f726e6("DB323_DM1_DM1{Nr}_bRoZB1", 2)
      ObjectEnable <- "DB322_DV1.DV1[Nr].bRoZB1"
      Appearance <- "DB323_DM1_DM1{Nr}_bRoZB1"
   Button "Button_15" at 820,677 size 97x35; TextOn 'OFF'; TextOff 'OFF'
      on Click: function_a9b64e44("DB323_DM1_DM1{Nr}_bRoZB1", 2)
      ObjectEnable <- "DB322_DV1.DV1[Nr].bRoZB1"
      Appearance <- "DB323_DM1_DM1{Nr}_bRoZB1"
   TextField "Text field_39" at 965,652 size 126x25; Text 'Wyjście steruj / Sterowanie'
   Circle "Circle_6" at 1012,680 size 30x30
      Appearance <- "DB323_DM1_DM1{Nr}_bWySter"
   Button "Button_16" at 29,687 size 188x32; TextOn 'Zawory i silniki'; TextOff 'DIO, AI, AO / Zawory i silniki'
      on Click: ActivateScreen("Service", 0)
*)